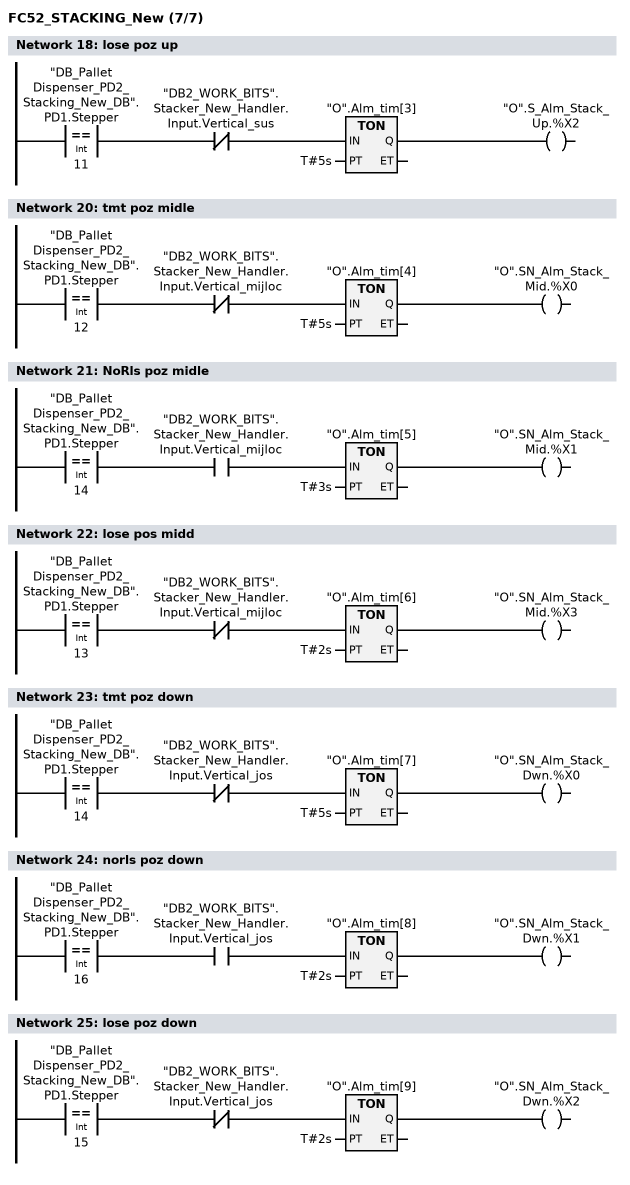
   "O".Alm_tim[3].TON(IN := ("DB_PalletDispenser_PD2_Stacking_New_DB".PD1.Stepper = 11) AND NOT "DB2_WORK_BITS".Stacker_New_Handler.Input.Vertical_sus,
                      PT := T#5s);
   "O".S_Alm_Stack_Up.%X2 := "O".Alm_tim[3].Q;
END_REGION

REGION Network 19: lose poz up
END_REGION

REGION Network 20: tmt poz midle
   "O".Alm_tim[4].TON(IN := ("DB_PalletDispenser_PD2_Stacking_New_DB".PD1.Stepper = 12) AND NOT "DB2_WORK_BITS".Stacker_New_Handler.Input.Vertical_mijloc,
                      PT := T#5s);
   "O".SN_Alm_Stack_Mid.%X0 := "O".Alm_tim[4].Q;
END_REGION

REGION Network 21: NoRls poz midle
   "O".Alm_tim[5].TON(IN := ("DB_PalletDispenser_PD2_Stacking_New_DB".PD1.Stepper = 14) AND "DB2_WORK_BITS".Stacker_New_Handler.Input.Vertical_mijloc,
                      PT := T#3s);
   "O".SN_Alm_Stack_Mid.%X1 := "O".Alm_tim[5].Q;
END_REGION

REGION Network 22: lose pos midd
   "O".Alm_tim[6].TON(IN := ("DB_PalletDispenser_PD2_Stacking_New_DB".PD1.Stepper = 13) AND NOT "DB2_WORK_BITS".Stacker_New_Handler.Input.Vertical_mijloc,
                      PT := T#2s);
   "O".SN_Alm_Stack_Mid.%X3 := "O".Alm_tim[6].Q;
END_REGION

REGION Network 23: tmt poz down
   "O".Alm_tim[7].TON(IN := ("DB_PalletDispenser_PD2_Stacking_New_DB".PD1.Stepper = 14) AND NOT "DB2_WORK_BITS".Stacker_New_Handler.Input.Vertical_jos,
                      PT := T#5s);
   "O".SN_Alm_Stack_Dwn.%X0 := "O".Alm_tim[7].Q;
END_REGION

REGION Network 24: norls poz down
   "O".Alm_tim[8].TON(IN := ("DB_PalletDispenser_PD2_Stacking_New_DB".PD1.Stepper = 16) AND "DB2_WORK_BITS".Stacker_New_Handler.Input.Vertical_jos,
                      PT := T#2s);
   "O".SN_Alm_Stack_Dwn.%X1 := "O".Alm_tim[8].Q;
END_REGION

REGION Network 25: lose poz down
   "O".Alm_tim[9].TON(IN := ("DB_PalletDispenser_PD2_Stacking_New_DB".PD1.Stepper = 15) AND NOT "DB2_WORK_BITS".Stacker_New_Handler.Input.Vertical_jos,
                      PT := T#2s);
   "O".SN_Alm_Stack_Dwn.%X2 := "O".Alm_tim[9].Q;
END_REGION
END_FUNCTION

FUNCTION "FC50_PALLET_LENGTH" : Void   // FC50, LAD
{ S7_Optimized_Access := 'TRUE' }
VERSION : 0.1
   VAR_INPUT
      Reset_counter_SN : Bool;
      Reset_counter_S : Bool;
   END_VAR
   VAR_TEMP
      Length1_UP : Bool;
   END_VAR
   VAR_TEMP   // added for the SCL form of the ladder/FBD networks
      _w1 : Bool;
   END_VAR
BEGIN

REGION Network 1
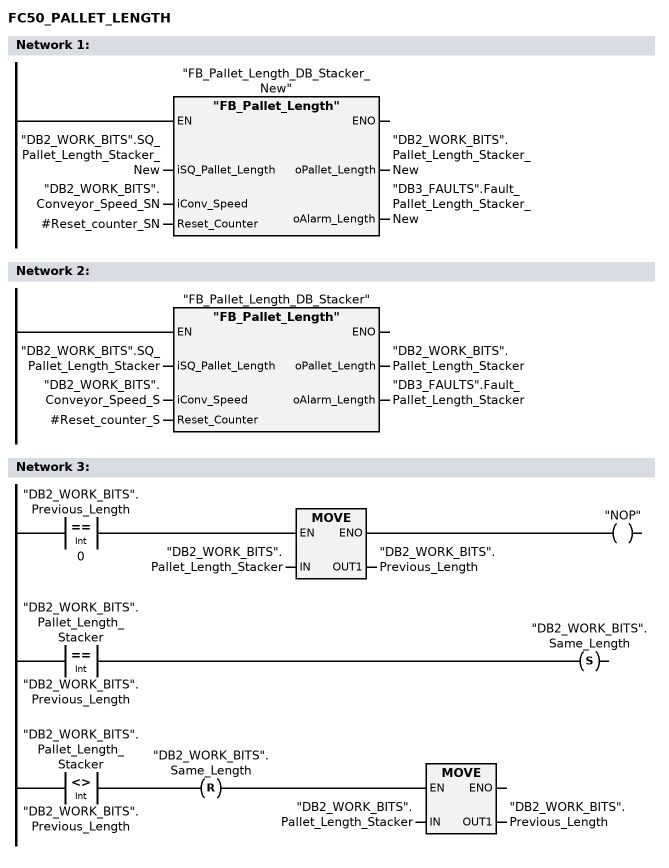
   RUNG wire#powerrail
      "FB_Pallet_Length_DB_Stacker_New"(iSQ_Pallet_Length := "DB2_WORK_BITS".SQ_Pallet_Length_Stacker_New, iConv_Speed := "DB2_WORK_BITS".Conveyor_Speed_SN, Reset_Counter := #Reset_counter_SN, oPallet_Length => "DB2_WORK_BITS".Pallet_Length_Stacker_New, oAlarm_Length => "DB3_FAULTS".Fault_Pallet_Length_Stacker_New)
   END_RUNG
   // the same network as SCL:
   "FB_Pallet_Length_DB_Stacker_New"(iSQ_Pallet_Length := "DB2_WORK_BITS".SQ_Pallet_Length_Stacker_New,   // "FB_Pallet_Length"
                           iConv_Speed := "DB2_WORK_BITS".Conveyor_Speed_SN,
                           Reset_Counter := #Reset_counter_SN,
                           oPallet_Length => "DB2_WORK_BITS".Pallet_Length_Stacker_New,
                           oAlarm_Length => "DB3_FAULTS".Fault_Pallet_Length_Stacker_New);
END_REGION

REGION Network 2
   RUNG wire#powerrail
      "FB_Pallet_Length_DB_Stacker"(iSQ_Pallet_Length := "DB2_WORK_BITS".SQ_Pallet_Length_Stacker, iConv_Speed := "DB2_WORK_BITS".Conveyor_Speed_S, Reset_Counter := #Reset_counter_S, oPallet_Length => "DB2_WORK_BITS".Pallet_Length_Stacker, oAlarm_Length => "DB3_FAULTS".Fault_Pallet_Length_Stacker)
   END_RUNG
   // the same network as SCL:
   "FB_Pallet_Length_DB_Stacker"(iSQ_Pallet_Length := "DB2_WORK_BITS".SQ_Pallet_Length_Stacker,   // "FB_Pallet_Length"
                           iConv_Speed := "DB2_WORK_BITS".Conveyor_Speed_S,
                           Reset_Counter := #Reset_counter_S,
                           oPallet_Length => "DB2_WORK_BITS".Pallet_Length_Stacker,
                           oAlarm_Length => "DB3_FAULTS".Fault_Pallet_Length_Stacker);
END_REGION

REGION Network 3
   RUNG wire#powerrail
      { S7_Templates := "SrcType := Int" } EQ_Contact(in1 := "DB2_WORK_BITS".Previous_Length, in2 := 0)
      Move(in := "DB2_WORK_BITS".Pallet_Length_Stacker, out1 => "DB2_WORK_BITS".Previous_Length)
      Coil( "NOP" )
   END_RUNG
   RUNG wire#powerrail
      { S7_Templates := "SrcType := Int" } EQ_Contact(in1 := "DB2_WORK_BITS".Pallet_Length_Stacker, in2 := "DB2_WORK_BITS".Previous_Length)
      S_Coil( "DB2_WORK_BITS".Same_Length )
   END_RUNG
   RUNG wire#powerrail
      { S7_Templates := "SrcType := Int" } NE_Contact(in1 := "DB2_WORK_BITS".Pallet_Length_Stacker, in2 := "DB2_WORK_BITS".Previous_Length)
      R_Coil( "DB2_WORK_BITS".Same_Length )
      Move(in := "DB2_WORK_BITS".Pallet_Length_Stacker, out1 => "DB2_WORK_BITS".Previous_Length)
   END_RUNG
   // the same network as SCL:
   #_w1 := "DB2_WORK_BITS".Previous_Length = 0;
   IF #_w1 THEN "DB2_WORK_BITS".Previous_Length := "DB2_WORK_BITS".Pallet_Length_Stacker; END_IF;
   "NOP" := #_w1;
   IF "DB2_WORK_BITS".Pallet_Length_Stacker = "DB2_WORK_BITS".Previous_Length THEN
       "DB2_WORK_BITS".Same_Length := TRUE;
   END_IF;
   IF "DB2_WORK_BITS".Pallet_Length_Stacker <> "DB2_WORK_BITS".Previous_Length THEN
       "DB2_WORK_BITS".Same_Length := FALSE;
       "DB2_WORK_BITS".Previous_Length := "DB2_WORK_BITS".Pallet_Length_Stacker;
   END_IF;
END_REGION
END_FUNCTION

FUNCTION "FC52_STACKING" : Void   // FC52, LAD
{ S7_Optimized_Access := 'TRUE' }
VERSION : 0.1
   VAR_TEMP
      Reset_S_Up : Bool;
      Reset_S_Fork : Bool;
      iB5_p : Bool;
      Reset_S : Bool;
      dumyb : Bool;
      dumyw : Int;
   END_VAR
   VAR_TEMP   // added for the SCL form of the ladder/FBD networks
      _w1 : Bool;
      _w2 : Bool;
      _w3 : Bool;
   END_VAR
BEGIN

REGION Network 1: mdm
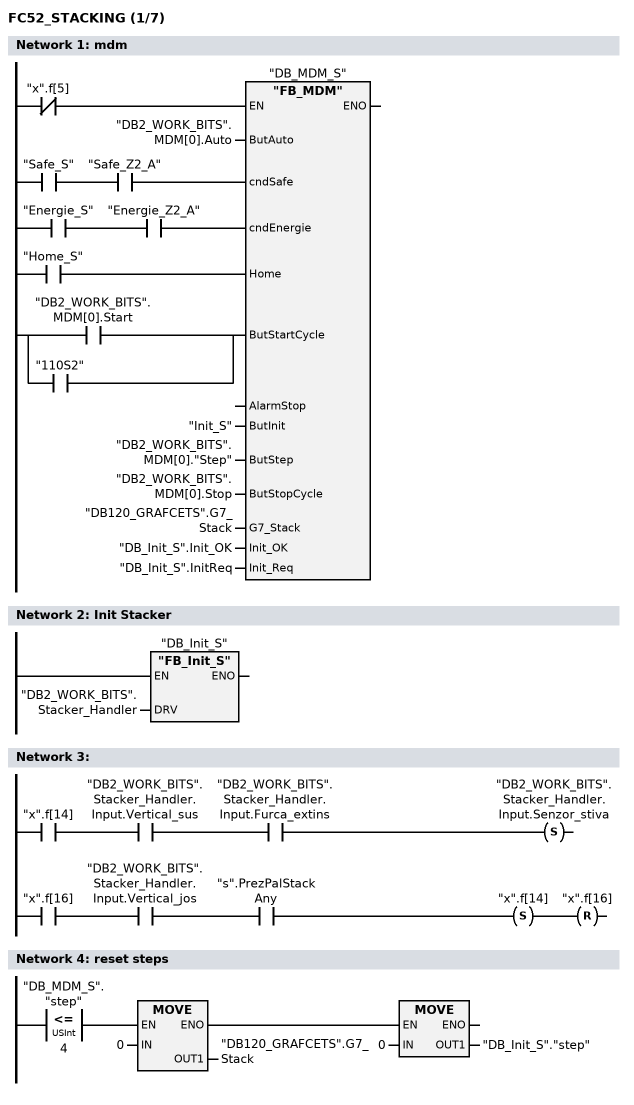
   RUNG wire#powerrail
      I_Contact( "x".f[5] )
      "DB_MDM_S"(cndSafe := wire#w1, cndEnergie := wire#w2, Home := wire#w3, ButStartCycle := wire#w4, ButAuto := "DB2_WORK_BITS".MDM[0].Auto, AlarmStop :=, ButInit := "Init_S", ButStep := "DB2_WORK_BITS".MDM[0]."Step", ButStopCycle := "DB2_WORK_BITS".MDM[0].Stop, G7_Stack := "DB120_GRAFCETS".G7_Stack, Init_OK := "DB_Init_S".Init_OK, Init_Req := "DB_Init_S".InitReq)
   END_RUNG
   RUNG wire#powerrail
      Contact( "Safe_S" )
      Contact( "Safe_Z2_A" )
   END_RUNG wire#w1
   RUNG wire#powerrail
      Contact( "Energie_S" )
      Contact( "Energie_Z2_A" )
   END_RUNG wire#w2
   RUNG wire#powerrail
      Contact( "Home_S" )
   END_RUNG wire#w3
   RUNG wire#powerrail
      Contact( "DB2_WORK_BITS".MDM[0].Start )
   END_RUNG wire#w4
   RUNG wire#powerrail
      Contact( "110S2" )
   END_RUNG wire#w4
   // the same network as SCL:
   IF NOT "x".f[5] THEN
       "DB_MDM_S"(ButAuto := "DB2_WORK_BITS".MDM[0].Auto,   // "FB_MDM"
                  cndSafe := "Safe_S" AND "Safe_Z2_A",
                  cndEnergie := "Energie_S" AND "Energie_Z2_A",
                  Home := "Home_S",
                  ButStartCycle := "DB2_WORK_BITS".MDM[0].Start OR "110S2",
                  ButInit := "Init_S",
                  ButStep := "DB2_WORK_BITS".MDM[0]."Step",
                  ButStopCycle := "DB2_WORK_BITS".MDM[0].Stop,
                  G7_Stack := "DB120_GRAFCETS".G7_Stack,
                  Init_OK := "DB_Init_S".Init_OK,
                  Init_Req := "DB_Init_S".InitReq);
   END_IF;
END_REGION

REGION Network 2: Init Stacker
   RUNG wire#powerrail
      "DB_Init_S"(DRV := "DB2_WORK_BITS".Stacker_Handler)
   END_RUNG
   // the same network as SCL:
   "DB_Init_S"(DRV := "DB2_WORK_BITS".Stacker_Handler);   // "FB_Init_S"
END_REGION

REGION Network 3
   RUNG wire#powerrail
      Contact( "x".f[14] )
      Contact( "DB2_WORK_BITS".Stacker_Handler.Input.Vertical_sus )
      Contact( "DB2_WORK_BITS".Stacker_Handler.Input.Furca_extins )
      S_Coil( "DB2_WORK_BITS".Stacker_Handler.Input.Senzor_stiva )
   END_RUNG
   RUNG wire#powerrail
      Contact( "x".f[16] )
      Contact( "DB2_WORK_BITS".Stacker_Handler.Input.Vertical_jos )
      Contact( "s".PrezPalStackAny )
      S_Coil( "x".f[14] )
      R_Coil( "x".f[16] )
   END_RUNG
   // the same network as SCL:
   IF "x".f[14] AND "DB2_WORK_BITS".Stacker_Handler.Input.Vertical_sus AND "DB2_WORK_BITS".Stacker_Handler.Input.Furca_extins THEN
       "DB2_WORK_BITS".Stacker_Handler.Input.Senzor_stiva := TRUE;
   END_IF;
   #_w1 := "x".f[16] AND "DB2_WORK_BITS".Stacker_Handler.Input.Vertical_jos AND "s".PrezPalStackAny;
   IF #_w1 THEN
       "x".f[14] := TRUE;
       "x".f[16] := FALSE;
   END_IF;
END_REGION

REGION Network 4: reset steps
   RUNG wire#powerrail
      { S7_Templates := "SrcType := USInt" } LE_Contact(in1 := "DB_MDM_S"."step", in2 := 4)
      Move(in := 0, out1 => "DB120_GRAFCETS".G7_Stack)
      Move(in := 0, out1 => "DB_Init_S"."step")
   END_RUNG
   // the same network as SCL:
   IF "DB_MDM_S"."step" <= 4 THEN
       "DB120_GRAFCETS".G7_Stack := 0;
       "DB_Init_S"."step" := 0;
   END_IF;
END_REGION

REGION Network 5: start graf stack
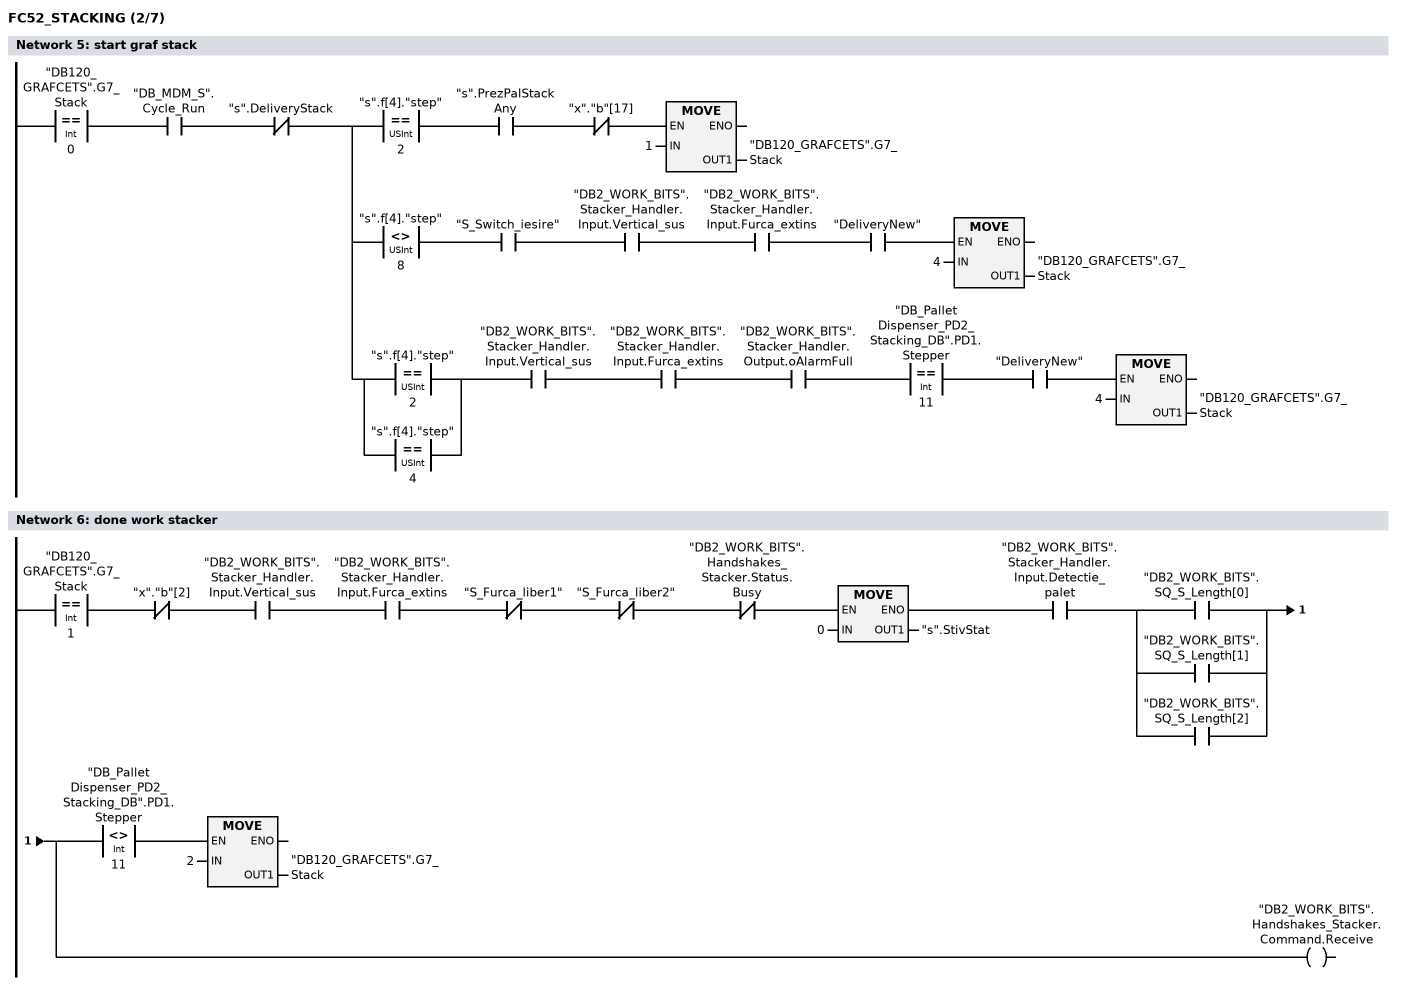
   RUNG wire#powerrail
      { S7_Templates := "SrcType := Int" } EQ_Contact(in1 := "DB120_GRAFCETS".G7_Stack, in2 := 0)
      Contact( "DB_MDM_S".Cycle_Run )
      I_Contact( "s".DeliveryStack )
      wire#w1
      { S7_Templates := "SrcType := USInt" } EQ_Contact(in1 := "s".f[4]."step", in2 := 2)
      Contact( "s".PrezPalStackAny )
      I_Contact( "x"."b"[17] )
      Move(in := 1, out1 => "DB120_GRAFCETS".G7_Stack)
   END_RUNG
   RUNG wire#w1
      { S7_Templates := "SrcType := USInt" } NE_Contact(in1 := "s".f[4]."step", in2 := 8)
      Contact( "S_Switch_iesire" )
      Contact( "DB2_WORK_BITS".Stacker_Handler.Input.Vertical_sus )
      Contact( "DB2_WORK_BITS".Stacker_Handler.Input.Furca_extins )
      Contact( "DeliveryNew" )
      Move(in := 4, out1 => "DB120_GRAFCETS".G7_Stack)
   END_RUNG
   RUNG wire#w1
      { S7_Templates := "SrcType := USInt" } EQ_Contact(in1 := "s".f[4]."step", in2 := 2)
      wire#w2
      Contact( "DB2_WORK_BITS".Stacker_Handler.Input.Vertical_sus )
      Contact( "DB2_WORK_BITS".Stacker_Handler.Input.Furca_extins )
      Contact( "DB2_WORK_BITS".Stacker_Handler.Output.oAlarmFull )
      { S7_Templates := "SrcType := Int" } EQ_Contact(in1 := "DB_PalletDispenser_PD2_Stacking_DB".PD1.Stepper, in2 := 11)
      Contact( "DeliveryNew" )
      Move(in := 4, out1 => "DB120_GRAFCETS".G7_Stack)
   END_RUNG
   RUNG wire#w1
      { S7_Templates := "SrcType := USInt" } EQ_Contact(in1 := "s".f[4]."step", in2 := 4)
   END_RUNG wire#w2
   // the same network as SCL:
   #_w1 := ("DB120_GRAFCETS".G7_Stack = 0) AND "DB_MDM_S".Cycle_Run AND NOT "s".DeliveryStack;
   IF #_w1 AND ("s".f[4]."step" = 2) AND "s".PrezPalStackAny AND NOT "x"."b"[17] THEN
       "DB120_GRAFCETS".G7_Stack := 1;
   END_IF;
   IF #_w1 AND ("s".f[4]."step" <> 8) AND "S_Switch_iesire" AND "DB2_WORK_BITS".Stacker_Handler.Input.Vertical_sus AND "DB2_WORK_BITS".Stacker_Handler.Input.Furca_extins AND "DeliveryNew" THEN
       "DB120_GRAFCETS".G7_Stack := 4;
   END_IF;
   IF #_w1 AND (("s".f[4]."step" = 2) OR ("s".f[4]."step" = 4)) AND "DB2_WORK_BITS".Stacker_Handler.Input.Vertical_sus AND "DB2_WORK_BITS".Stacker_Handler.Input.Furca_extins AND "DB2_WORK_BITS".Stacker_Handler.Output.oAlarmFull AND ("DB_PalletDispenser_PD2_Stacking_DB".PD1.Stepper = 11) AND "DeliveryNew" THEN
       "DB120_GRAFCETS".G7_Stack := 4;
   END_IF;
END_REGION

REGION Network 6: done work stacker
   RUNG wire#powerrail
      { S7_Templates := "SrcType := Int" } EQ_Contact(in1 := "DB120_GRAFCETS".G7_Stack, in2 := 1)
      I_Contact( "x"."b"[2] )
      Contact( "DB2_WORK_BITS".Stacker_Handler.Input.Vertical_sus )
      Contact( "DB2_WORK_BITS".Stacker_Handler.Input.Furca_extins )
      I_Contact( "S_Furca_liber1" )
      I_Contact( "S_Furca_liber2" )
      I_Contact( "DB2_WORK_BITS".Handshakes_Stacker.Status.Busy )
      Move(in := 0, out1 => "s".StivStat)
      Contact( "DB2_WORK_BITS".Stacker_Handler.Input.Detectie_palet )
      wire#w1
      Contact( "DB2_WORK_BITS".SQ_S_Length[0] )
      wire#w2
      { S7_Templates := "SrcType := Int" } NE_Contact(in1 := "DB_PalletDispenser_PD2_Stacking_DB".PD1.Stepper, in2 := 11)
      Move(in := 2, out1 => "DB120_GRAFCETS".G7_Stack)
   END_RUNG
   RUNG wire#w1
      Contact( "DB2_WORK_BITS".SQ_S_Length[1] )
   END_RUNG wire#w2
   RUNG wire#w1
      Contact( "DB2_WORK_BITS".SQ_S_Length[2] )
   END_RUNG wire#w2
   RUNG wire#w2
      Coil( "DB2_WORK_BITS".Handshakes_Stacker.Command.Receive )
   END_RUNG
   // the same network as SCL:
   #_w1 := ("DB120_GRAFCETS".G7_Stack = 1) AND NOT "x"."b"[2] AND "DB2_WORK_BITS".Stacker_Handler.Input.Vertical_sus AND "DB2_WORK_BITS".Stacker_Handler.Input.Furca_extins AND NOT "S_Furca_liber1" AND NOT "S_Furca_liber2" AND NOT "DB2_WORK_BITS".Handshakes_Stacker.Status.Busy;
   IF #_w1 THEN "s".StivStat := 0; END_IF;
   #_w2 := #_w1 AND "DB2_WORK_BITS".Stacker_Handler.Input.Detectie_palet AND ("DB2_WORK_BITS".SQ_S_Length[0] OR "DB2_WORK_BITS".SQ_S_Length[1] OR "DB2_WORK_BITS".SQ_S_Length[2]);
   IF #_w2 AND ("DB_PalletDispenser_PD2_Stacking_DB".PD1.Stepper <> 11) THEN
       "DB120_GRAFCETS".G7_Stack := 2;
   END_IF;
   "DB2_WORK_BITS".Handshakes_Stacker.Command.Receive := #_w2;
END_REGION

REGION Network 7: decision continue/release stack
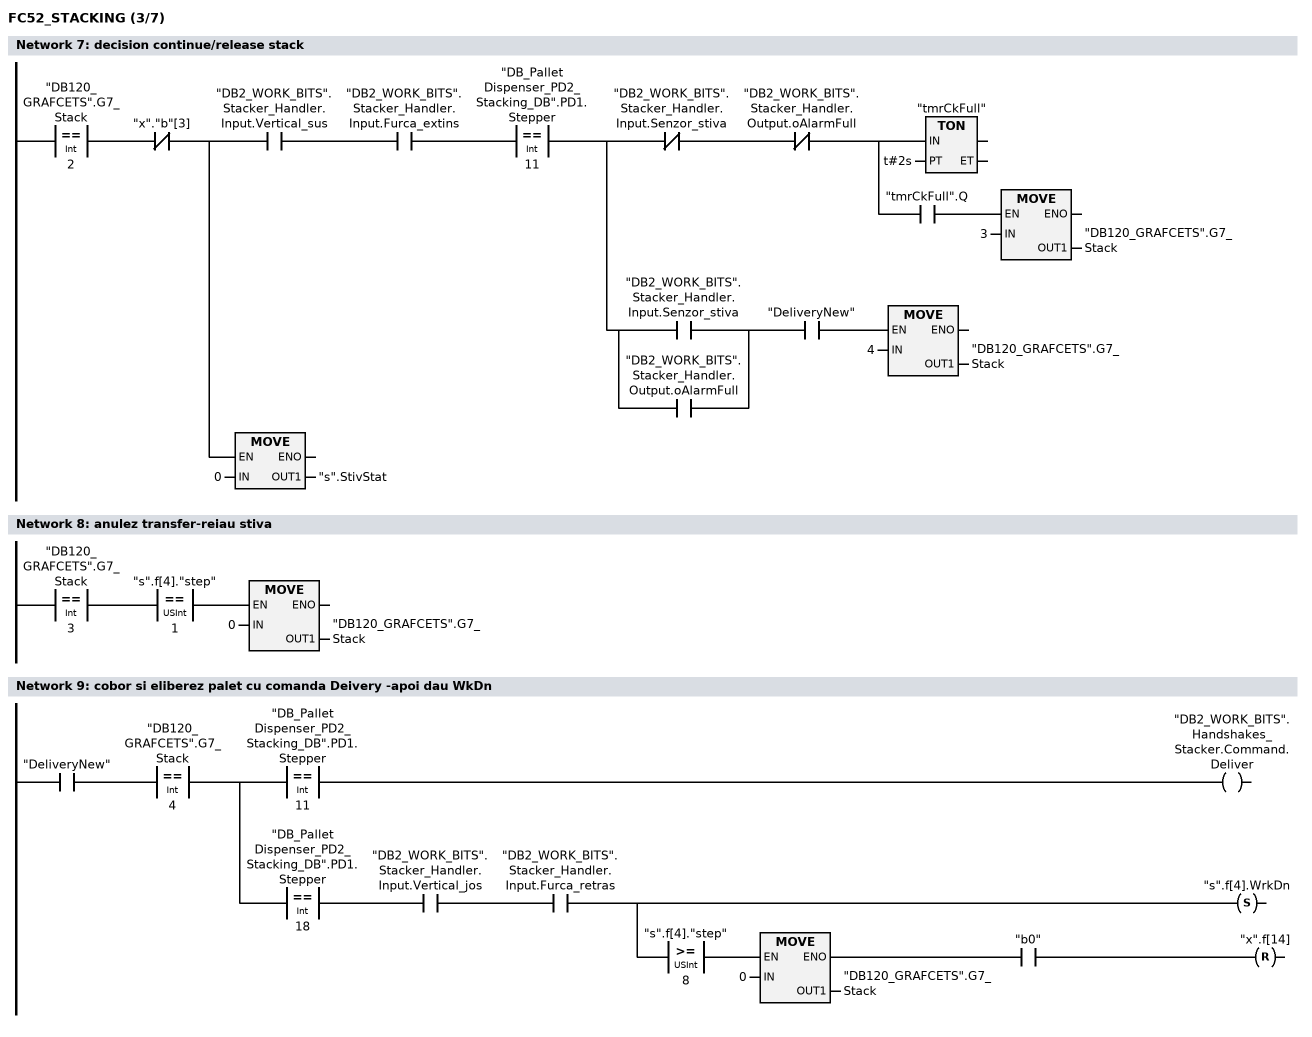
   #_w1 := ("DB120_GRAFCETS".G7_Stack = 2) AND NOT "x"."b"[3];
   #_w2 := #_w1 AND "DB2_WORK_BITS".Stacker_Handler.Input.Vertical_sus AND "DB2_WORK_BITS".Stacker_Handler.Input.Furca_extins AND ("DB_PalletDispenser_PD2_Stacking_DB".PD1.Stepper = 11);
   #_w3 := #_w2 AND NOT "DB2_WORK_BITS".Stacker_Handler.Input.Senzor_stiva AND NOT "DB2_WORK_BITS".Stacker_Handler.Output.oAlarmFull;
   "tmrCkFull".TON(IN := #_w3, PT := t#2s);
   IF #_w3 AND "tmrCkFull".Q THEN "DB120_GRAFCETS".G7_Stack := 3; END_IF;
   IF #_w2 AND ("DB2_WORK_BITS".Stacker_Handler.Input.Senzor_stiva OR "DB2_WORK_BITS".Stacker_Handler.Output.oAlarmFull) AND "DeliveryNew" THEN
       "DB120_GRAFCETS".G7_Stack := 4;
   END_IF;
   IF #_w1 THEN "s".StivStat := 0; END_IF;
END_REGION

REGION Network 8: anulez transfer-reiau stiva
   RUNG wire#powerrail
      { S7_Templates := "SrcType := Int" } EQ_Contact(in1 := "DB120_GRAFCETS".G7_Stack, in2 := 3)
      { S7_Templates := "SrcType := USInt" } EQ_Contact(in1 := "s".f[4]."step", in2 := 1)
      Move(in := 0, out1 => "DB120_GRAFCETS".G7_Stack)
   END_RUNG
   // the same network as SCL:
   IF ("DB120_GRAFCETS".G7_Stack = 3) AND ("s".f[4]."step" = 1) THEN "DB120_GRAFCETS".G7_Stack := 0; END_IF;
END_REGION

REGION Network 9: cobor si eliberez palet cu comanda Deivery -apoi dau WkDn
   RUNG wire#powerrail
      Contact( "DeliveryNew" )
      { S7_Templates := "SrcType := Int" } EQ_Contact(in1 := "DB120_GRAFCETS".G7_Stack, in2 := 4)
      wire#w1
      { S7_Templates := "SrcType := Int" } EQ_Contact(in1 := "DB_PalletDispenser_PD2_Stacking_DB".PD1.Stepper, in2 := 11)
      Coil( "DB2_WORK_BITS".Handshakes_Stacker.Command.Deliver )
   END_RUNG
   RUNG wire#w1
      { S7_Templates := "SrcType := Int" } EQ_Contact(in1 := "DB_PalletDispenser_PD2_Stacking_DB".PD1.Stepper, in2 := 18)
      Contact( "DB2_WORK_BITS".Stacker_Handler.Input.Vertical_jos )
      Contact( "DB2_WORK_BITS".Stacker_Handler.Input.Furca_retras )
      wire#w2
      S_Coil( "s".f[4].WrkDn )
   END_RUNG
   RUNG wire#w2
      { S7_Templates := "SrcType := USInt" } GE_Contact(in1 := "s".f[4]."step", in2 := 8)
      Move(in := 0, out1 => "DB120_GRAFCETS".G7_Stack)
      Contact( "b0" )
      R_Coil( "x".f[14] )
   END_RUNG
   // the same network as SCL:
   #_w1 := "DeliveryNew" AND ("DB120_GRAFCETS".G7_Stack = 4);
   "DB2_WORK_BITS".Handshakes_Stacker.Command.Deliver := #_w1 AND ("DB_PalletDispenser_PD2_Stacking_DB".PD1.Stepper = 11);
   #_w2 := #_w1 AND ("DB_PalletDispenser_PD2_Stacking_DB".PD1.Stepper = 18) AND "DB2_WORK_BITS".Stacker_Handler.Input.Vertical_jos AND "DB2_WORK_BITS".Stacker_Handler.Input.Furca_retras;
   IF #_w2 THEN "s".f[4].WrkDn := TRUE; END_IF;
   #_w3 := #_w2 AND ("s".f[4]."step" >= 8);
   IF #_w3 THEN "DB120_GRAFCETS".G7_Stack := 0; END_IF;
   IF #_w3 AND "b0" THEN "x".f[14] := FALSE; END_IF;
END_REGION

REGION Network 10: delivery
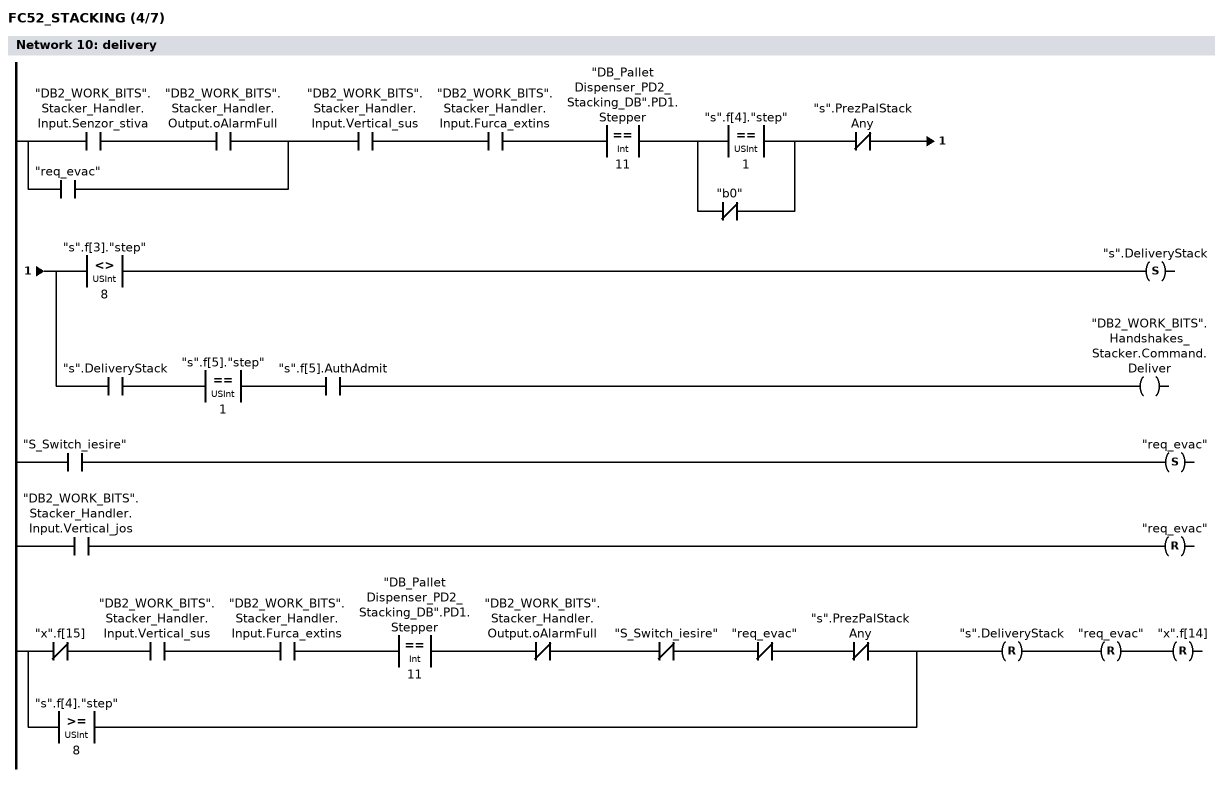
   RUNG wire#powerrail
      Contact( "DB2_WORK_BITS".Stacker_Handler.Input.Senzor_stiva )
      Contact( "DB2_WORK_BITS".Stacker_Handler.Output.oAlarmFull )
      wire#w1
      Contact( "DB2_WORK_BITS".Stacker_Handler.Input.Vertical_sus )
      Contact( "DB2_WORK_BITS".Stacker_Handler.Input.Furca_extins )
      { S7_Templates := "SrcType := Int" } EQ_Contact(in1 := "DB_PalletDispenser_PD2_Stacking_DB".PD1.Stepper, in2 := 11)
      wire#w2
      { S7_Templates := "SrcType := USInt" } EQ_Contact(in1 := "s".f[4]."step", in2 := 1)
      wire#w3
      I_Contact( "s".PrezPalStackAny )
      wire#w4
      { S7_Templates := "SrcType := USInt" } NE_Contact(in1 := "s".f[3]."step", in2 := 8)
      S_Coil( "s".DeliveryStack )
   END_RUNG
   RUNG wire#powerrail
      Contact( "req_evac" )
   END_RUNG wire#w1
   RUNG wire#w2
      I_Contact( "b0" )
   END_RUNG wire#w3
   RUNG wire#w4
      Contact( "s".DeliveryStack )
      { S7_Templates := "SrcType := USInt" } EQ_Contact(in1 := "s".f[5]."step", in2 := 1)
      Contact( "s".f[5].AuthAdmit )
      Coil( "DB2_WORK_BITS".Handshakes_Stacker.Command.Deliver )
   END_RUNG
   RUNG wire#powerrail
      Contact( "S_Switch_iesire" )
      S_Coil( "req_evac" )
   END_RUNG
   RUNG wire#powerrail
      Contact( "DB2_WORK_BITS".Stacker_Handler.Input.Vertical_jos )
      R_Coil( "req_evac" )
   END_RUNG
   RUNG wire#powerrail
      I_Contact( "x".f[15] )
      Contact( "DB2_WORK_BITS".Stacker_Handler.Input.Vertical_sus )
      Contact( "DB2_WORK_BITS".Stacker_Handler.Input.Furca_extins )
      { S7_Templates := "SrcType := Int" } EQ_Contact(in1 := "DB_PalletDispenser_PD2_Stacking_DB".PD1.Stepper, in2 := 11)
      I_Contact( "DB2_WORK_BITS".Stacker_Handler.Output.oAlarmFull )
      I_Contact( "S_Switch_iesire" )
      I_Contact( "req_evac" )
      I_Contact( "s".PrezPalStackAny )
      wire#w5
      R_Coil( "s".DeliveryStack )
      R_Coil( "req_evac" )
      R_Coil( "x".f[14] )
   END_RUNG
   RUNG wire#powerrail
      { S7_Templates := "SrcType := USInt" } GE_Contact(in1 := "s".f[4]."step", in2 := 8)
   END_RUNG wire#w5
   // the same network as SCL:
   #_w1 := (("DB2_WORK_BITS".Stacker_Handler.Input.Senzor_stiva AND "DB2_WORK_BITS".Stacker_Handler.Output.oAlarmFull) OR "req_evac") AND "DB2_WORK_BITS".Stacker_Handler.Input.Vertical_sus AND "DB2_WORK_BITS".Stacker_Handler.Input.Furca_extins AND ("DB_PalletDispenser_PD2_Stacking_DB".PD1.Stepper = 11) AND (("s".f[4]."step" = 1) OR NOT "b0") AND NOT "s".PrezPalStackAny;
   IF #_w1 AND ("s".f[3]."step" <> 8) THEN "s".DeliveryStack := TRUE; END_IF;
   "DB2_WORK_BITS".Handshakes_Stacker.Command.Deliver := #_w1 AND "s".DeliveryStack AND ("s".f[5]."step" = 1) AND "s".f[5].AuthAdmit;
   IF "S_Switch_iesire" THEN "req_evac" := TRUE; END_IF;
   IF "DB2_WORK_BITS".Stacker_Handler.Input.Vertical_jos THEN "req_evac" := FALSE; END_IF;
   IF (NOT "x".f[15] AND "DB2_WORK_BITS".Stacker_Handler.Input.Vertical_sus AND "DB2_WORK_BITS".Stacker_Handler.Input.Furca_extins AND ("DB_PalletDispenser_PD2_Stacking_DB".PD1.Stepper = 11) AND NOT "DB2_WORK_BITS".Stacker_Handler.Output.oAlarmFull AND NOT "S_Switch_iesire" AND NOT "req_evac" AND NOT "s".PrezPalStackAny) OR ("s".f[4]."step" >= 8) THEN
       "s".DeliveryStack := FALSE;
   END_IF;
   #_w2 := (NOT "x".f[15] AND "DB2_WORK_BITS".Stacker_Handler.Input.Vertical_sus AND "DB2_WORK_BITS".Stacker_Handler.Input.Furca_extins AND ("DB_PalletDispenser_PD2_Stacking_DB".PD1.Stepper = 11) AND NOT "DB2_WORK_BITS".Stacker_Handler.Output.oAlarmFull AND NOT "S_Switch_iesire" AND NOT "req_evac" AND NOT "s".PrezPalStackAny) OR ("s".f[4]."step" >= 8);
   IF #_w2 THEN
       "req_evac" := FALSE;
       "x".f[14] := FALSE;
   END_IF;
END_REGION

REGION Network 11: call FB stack
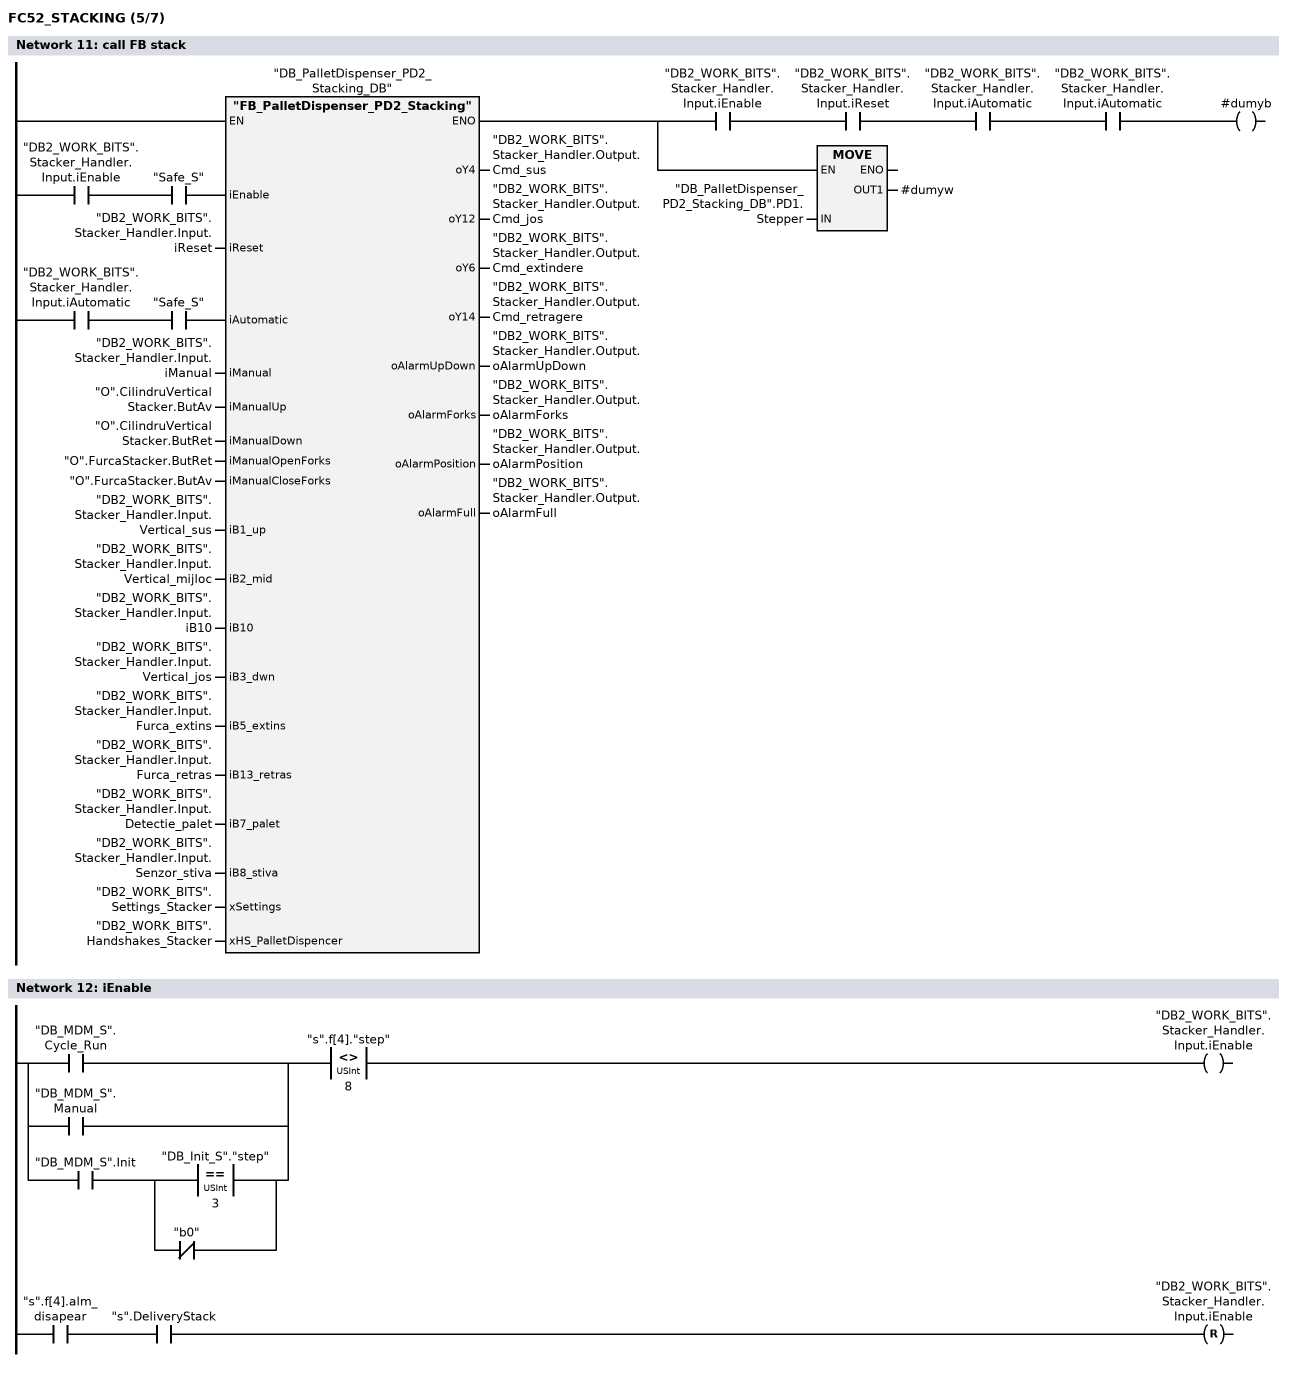
   RUNG wire#powerrail
      "DB_PalletDispenser_PD2_Stacking_DB"(iEnable := wire#w1, iAutomatic := wire#w2, iReset := "DB2_WORK_BITS".Stacker_Handler.Input.iReset, iManual := "DB2_WORK_BITS".Stacker_Handler.Input.iManual, iManualUp := "O".CilindruVerticalStacker.ButAv, iManualDown := "O".CilindruVerticalStacker.ButRet, iManualOpenForks := "O".FurcaStacker.ButRet, iManualCloseForks := "O".FurcaStacker.ButAv, iB1_up := "DB2_WORK_BITS".Stacker_Handler.Input.Vertical_sus, iB2_mid := "DB2_WORK_BITS".Stacker_Handler.Input.Vertical_mijloc, iB10 := "DB2_WORK_BITS".Stacker_Handler.Input.iB10, iB3_dwn := "DB2_WORK_BITS".Stacker_Handler.Input.Vertical_jos, iB5_extins := "DB2_WORK_BITS".Stacker_Handler.Input.Furca_extins, iB13_retras := "DB2_WORK_BITS".Stacker_Handler.Input.Furca_retras, iB7_palet := "DB2_WORK_BITS".Stacker_Handler.Input.Detectie_palet, iB8_stiva := "DB2_WORK_BITS".Stacker_Handler.Input.Senzor_stiva, xSettings := "DB2_WORK_BITS".Settings_Stacker, xHS_PalletDispencer := "DB2_WORK_BITS".Handshakes_Stacker, oY4 => "DB2_WORK_BITS".Stacker_Handler.Output.Cmd_sus, oY12 => "DB2_WORK_BITS".Stacker_Handler.Output.Cmd_jos, oY6 => "DB2_WORK_BITS".Stacker_Handler.Output.Cmd_extindere, oY14 => "DB2_WORK_BITS".Stacker_Handler.Output.Cmd_retragere, oAlarmUpDown => "DB2_WORK_BITS".Stacker_Handler.Output.oAlarmUpDown, oAlarmForks => "DB2_WORK_BITS".Stacker_Handler.Output.oAlarmForks, oAlarmPosition => "DB2_WORK_BITS".Stacker_Handler.Output.oAlarmPosition, oAlarmFull => "DB2_WORK_BITS".Stacker_Handler.Output.oAlarmFull)
      wire#w3
      Contact( "DB2_WORK_BITS".Stacker_Handler.Input.iEnable )
      Contact( "DB2_WORK_BITS".Stacker_Handler.Input.iReset )
      Contact( "DB2_WORK_BITS".Stacker_Handler.Input.iAutomatic )
      Contact( "DB2_WORK_BITS".Stacker_Handler.Input.iAutomatic )
      Coil( #dumyb )
   END_RUNG
   RUNG wire#powerrail
      Contact( "DB2_WORK_BITS".Stacker_Handler.Input.iEnable )
      Contact( "Safe_S" )
   END_RUNG wire#w1
   RUNG wire#powerrail
      Contact( "DB2_WORK_BITS".Stacker_Handler.Input.iAutomatic )
      Contact( "Safe_S" )
   END_RUNG wire#w2
   RUNG wire#w3
      Move(in := "DB_PalletDispenser_PD2_Stacking_DB".PD1.Stepper, out1 => #dumyw)
   END_RUNG
   // the same network as SCL:
   "DB_PalletDispenser_PD2_Stacking_DB"(iEnable := "DB2_WORK_BITS".Stacker_Handler.Input.iEnable AND "Safe_S",   // "FB_PalletDispenser_PD2_Stacking"